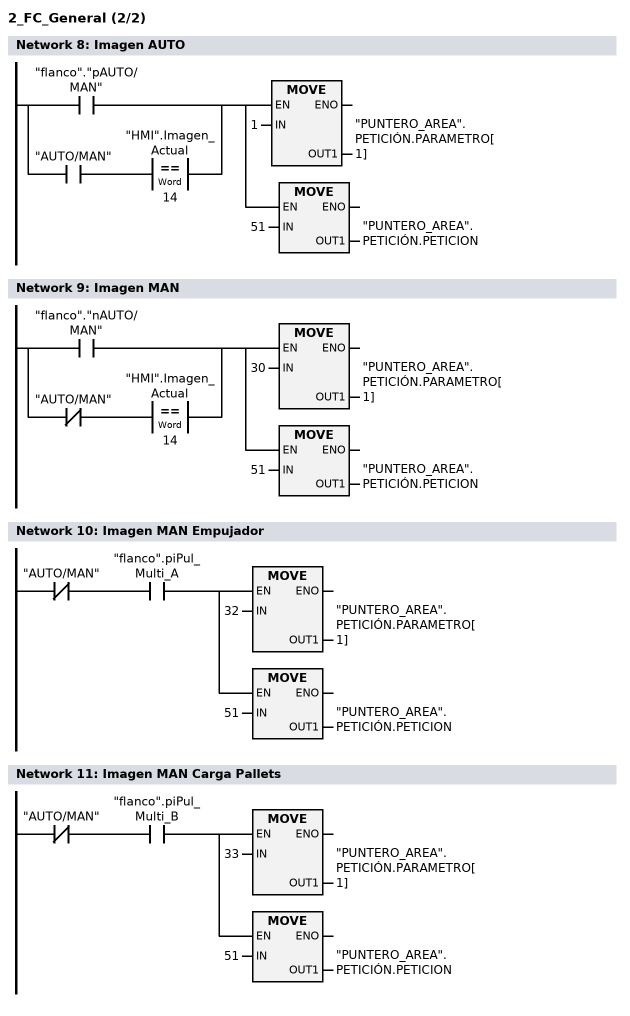
   RUNG wire#powerrail
      Contact( "flanco"."pAUTO/MAN" )
      wire#w1
      { S7_GenerateENO := "TRUE" } Move(in := 1, out1 => "PUNTERO_AREA".PETICIÓN.PARAMETRO[1])
   END_RUNG
   RUNG wire#powerrail
      Contact( "AUTO/MAN" )
      { S7_Templates := "SrcType := Word" } EQ_Contact(in1 := "HMI".Imagen_Actual, in2 := 14)
   END_RUNG wire#w1
   RUNG wire#w1
      { S7_GenerateENO := "TRUE" } Move(in := 51, out1 => "PUNTERO_AREA".PETICIÓN.PETICION)
   END_RUNG
   // the same network as SCL:
   IF "flanco"."pAUTO/MAN" OR ("AUTO/MAN" AND ("HMI".Imagen_Actual = 14)) THEN
       "PUNTERO_AREA".PETICIÓN.PARAMETRO[1] := 1;
       "PUNTERO_AREA".PETICIÓN.PETICION := 51;
   END_IF;
END_REGION

REGION Network 9: Imagen MAN
   RUNG wire#powerrail
      Contact( "flanco"."nAUTO/MAN" )
      wire#w1
      { S7_GenerateENO := "TRUE" } Move(in := 30, out1 => "PUNTERO_AREA".PETICIÓN.PARAMETRO[1])
   END_RUNG
   RUNG wire#powerrail
      I_Contact( "AUTO/MAN" )
      { S7_Templates := "SrcType := Word" } EQ_Contact(in1 := "HMI".Imagen_Actual, in2 := 14)
   END_RUNG wire#w1
   RUNG wire#w1
      { S7_GenerateENO := "TRUE" } Move(in := 51, out1 => "PUNTERO_AREA".PETICIÓN.PETICION)
   END_RUNG
   // the same network as SCL:
   IF "flanco"."nAUTO/MAN" OR (NOT "AUTO/MAN" AND ("HMI".Imagen_Actual = 14)) THEN
       "PUNTERO_AREA".PETICIÓN.PARAMETRO[1] := 30;
       "PUNTERO_AREA".PETICIÓN.PETICION := 51;
   END_IF;
END_REGION

REGION Network 10: Imagen MAN Empujador
   RUNG wire#powerrail
      I_Contact( "AUTO/MAN" )
      Contact( "flanco".piPul_Multi_A )
      wire#w1
      { S7_GenerateENO := "TRUE" } Move(in := 32, out1 => "PUNTERO_AREA".PETICIÓN.PARAMETRO[1])
   END_RUNG
   RUNG wire#w1
      { S7_GenerateENO := "TRUE" } Move(in := 51, out1 => "PUNTERO_AREA".PETICIÓN.PETICION)
   END_RUNG
   // the same network as SCL:
   IF NOT "AUTO/MAN" AND "flanco".piPul_Multi_A THEN
       "PUNTERO_AREA".PETICIÓN.PARAMETRO[1] := 32;
       "PUNTERO_AREA".PETICIÓN.PETICION := 51;
   END_IF;
END_REGION

REGION Network 11: Imagen MAN Carga Pallets
   RUNG wire#powerrail
      I_Contact( "AUTO/MAN" )
      Contact( "flanco".piPul_Multi_B )
      wire#w1
      { S7_GenerateENO := "TRUE" } Move(in := 33, out1 => "PUNTERO_AREA".PETICIÓN.PARAMETRO[1])
   END_RUNG
   RUNG wire#w1
      { S7_GenerateENO := "TRUE" } Move(in := 51, out1 => "PUNTERO_AREA".PETICIÓN.PETICION)
   END_RUNG
   // the same network as SCL:
   IF NOT "AUTO/MAN" AND "flanco".piPul_Multi_B THEN
       "PUNTERO_AREA".PETICIÓN.PARAMETRO[1] := 33;
       "PUNTERO_AREA".PETICIÓN.PETICION := 51;
   END_IF;
END_REGION
END_FUNCTION

FUNCTION "1_FC_Inv_Entradas" : Void   // FC9, LAD
{ S7_Optimized_Access := 'FALSE' }
VERSION : 0.1
BEGIN

REGION Network 1: "iiPul_DeshCargPall"
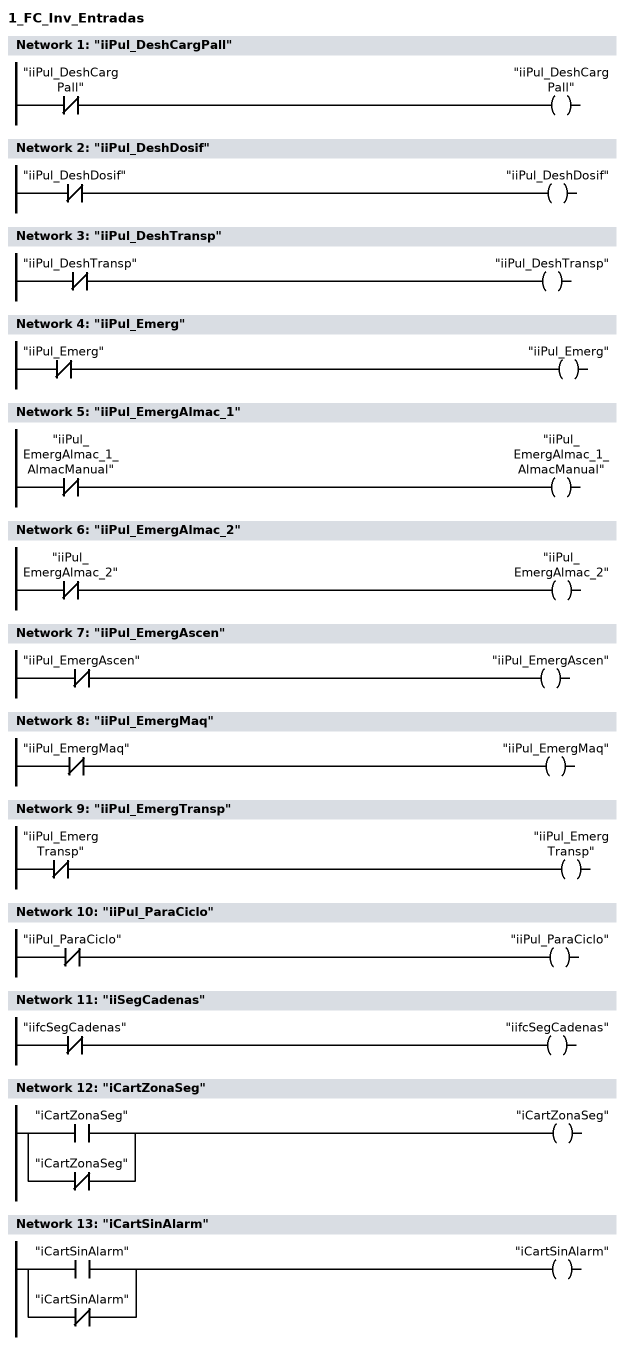
   RUNG wire#powerrail
      I_Contact( "iiPul_DeshCargPall" )
      Coil( "iiPul_DeshCargPall" )
   END_RUNG
   // the same network as SCL:
   "iiPul_DeshCargPall" := NOT "iiPul_DeshCargPall";
END_REGION

REGION Network 2: "iiPul_DeshDosif"
   RUNG wire#powerrail
      I_Contact( "iiPul_DeshDosif" )
      Coil( "iiPul_DeshDosif" )
   END_RUNG
   // the same network as SCL:
   "iiPul_DeshDosif" := NOT "iiPul_DeshDosif";
END_REGION

REGION Network 3: "iiPul_DeshTransp"
   RUNG wire#powerrail
      I_Contact( "iiPul_DeshTransp" )
      Coil( "iiPul_DeshTransp" )
   END_RUNG
   // the same network as SCL:
   "iiPul_DeshTransp" := NOT "iiPul_DeshTransp";
END_REGION

REGION Network 4: "iiPul_Emerg"
   RUNG wire#powerrail
      I_Contact( "iiPul_Emerg" )
      Coil( "iiPul_Emerg" )
   END_RUNG
   // the same network as SCL:
   "iiPul_Emerg" := NOT "iiPul_Emerg";
END_REGION

REGION Network 5: "iiPul_EmergAlmac_1"
   RUNG wire#powerrail
      I_Contact( "iiPul_EmergAlmac_1_AlmacManual" )
      Coil( "iiPul_EmergAlmac_1_AlmacManual" )
   END_RUNG
   // the same network as SCL:
   "iiPul_EmergAlmac_1_AlmacManual" := NOT "iiPul_EmergAlmac_1_AlmacManual";
END_REGION

REGION Network 6: "iiPul_EmergAlmac_2"
   RUNG wire#powerrail
      I_Contact( "iiPul_EmergAlmac_2" )
      Coil( "iiPul_EmergAlmac_2" )
   END_RUNG
   // the same network as SCL:
   "iiPul_EmergAlmac_2" := NOT "iiPul_EmergAlmac_2";
END_REGION

REGION Network 7: "iiPul_EmergAscen"
   RUNG wire#powerrail
      I_Contact( "iiPul_EmergAscen" )
      Coil( "iiPul_EmergAscen" )
   END_RUNG
   // the same network as SCL:
   "iiPul_EmergAscen" := NOT "iiPul_EmergAscen";
END_REGION

REGION Network 8: "iiPul_EmergMaq"
   RUNG wire#powerrail
      I_Contact( "iiPul_EmergMaq" )
      Coil( "iiPul_EmergMaq" )
   END_RUNG
   // the same network as SCL:
   "iiPul_EmergMaq" := NOT "iiPul_EmergMaq";
END_REGION

REGION Network 9: "iiPul_EmergTransp"
   RUNG wire#powerrail
      I_Contact( "iiPul_EmergTransp" )
      Coil( "iiPul_EmergTransp" )
   END_RUNG
   // the same network as SCL:
   "iiPul_EmergTransp" := NOT "iiPul_EmergTransp";
END_REGION

REGION Network 10: "iiPul_ParaCiclo"
   RUNG wire#powerrail
      I_Contact( "iiPul_ParaCiclo" )
      Coil( "iiPul_ParaCiclo" )
   END_RUNG
   // the same network as SCL:
   "iiPul_ParaCiclo" := NOT "iiPul_ParaCiclo";
END_REGION

REGION Network 11: "iiSegCadenas"
   RUNG wire#powerrail
      I_Contact( "iifcSegCadenas" )
      Coil( "iifcSegCadenas" )
   END_RUNG
   // the same network as SCL:
   "iifcSegCadenas" := NOT "iifcSegCadenas";
END_REGION

REGION Network 12: "iCartZonaSeg"
   RUNG wire#powerrail
      Contact( "iCartZonaSeg" )
      wire#w1
      Coil( "iCartZonaSeg" )
   END_RUNG
   RUNG wire#powerrail
      I_Contact( "iCartZonaSeg" )
   END_RUNG wire#w1
   // the same network as SCL:
   "iCartZonaSeg" := "iCartZonaSeg" OR NOT "iCartZonaSeg";
END_REGION

REGION Network 13: "iCartSinAlarm"
   RUNG wire#powerrail
      Contact( "iCartSinAlarm" )
      wire#w1
      Coil( "iCartSinAlarm" )
   END_RUNG
   RUNG wire#powerrail
      I_Contact( "iCartSinAlarm" )
   END_RUNG wire#w1
   // the same network as SCL:
   "iCartSinAlarm" := "iCartSinAlarm" OR NOT "iCartSinAlarm";
END_REGION
END_FUNCTION

FUNCTION "9_FC_Salidas" : Void   // FC10, LAD
{ S7_Optimized_Access := 'FALSE' }
VERSION : 0.1
BEGIN

REGION Network 1: "oLuz_CicloHab"
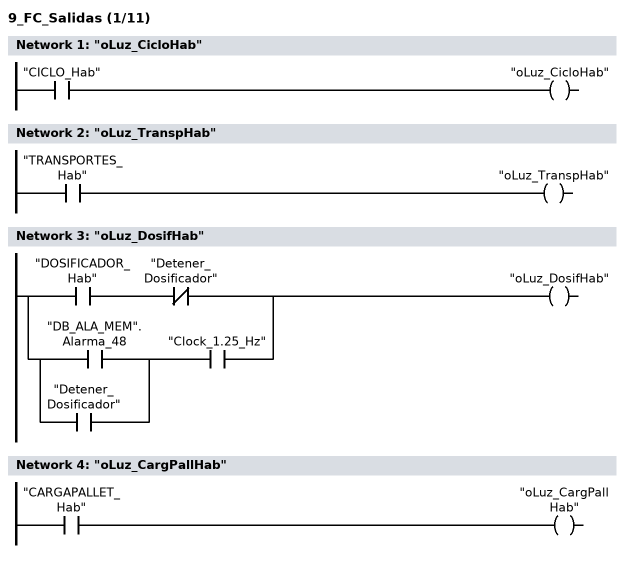
   RUNG wire#powerrail
      Contact( "CICLO_Hab" )
      Coil( "oLuz_CicloHab" )
   END_RUNG
   // the same network as SCL:
   "oLuz_CicloHab" := "CICLO_Hab";
END_REGION

REGION Network 2: "oLuz_TranspHab"
   RUNG wire#powerrail
      Contact( "TRANSPORTES_Hab" )
      Coil( "oLuz_TranspHab" )
   END_RUNG
   // the same network as SCL:
   "oLuz_TranspHab" := "TRANSPORTES_Hab";
END_REGION

REGION Network 3: "oLuz_DosifHab"
   RUNG wire#powerrail
      Contact( "DOSIFICADOR_Hab" )
      I_Contact( "Detener_Dosificador" )
      wire#w1
      Coil( "oLuz_DosifHab" )
   END_RUNG
   RUNG wire#powerrail
      Contact( "DB_ALA_MEM".Alarma_48 )
      wire#w2
      Contact( "Clock_1.25_Hz" )
   END_RUNG wire#w1
   RUNG wire#powerrail
      Contact( "Detener_Dosificador" )
   END_RUNG wire#w2
   // the same network as SCL:
   "oLuz_DosifHab" := ("DOSIFICADOR_Hab" AND NOT "Detener_Dosificador") OR (("DB_ALA_MEM".Alarma_48 OR "Detener_Dosificador") AND "Clock_1.25_Hz");
END_REGION

REGION Network 4: "oLuz_CargPallHab"
   RUNG wire#powerrail
      Contact( "CARGAPALLET_Hab" )
      Coil( "oLuz_CargPallHab" )
   END_RUNG
   // the same network as SCL:
   "oLuz_CargPallHab" := "CARGAPALLET_Hab";
END_REGION

REGION Network 5: "oLuz_Segur"
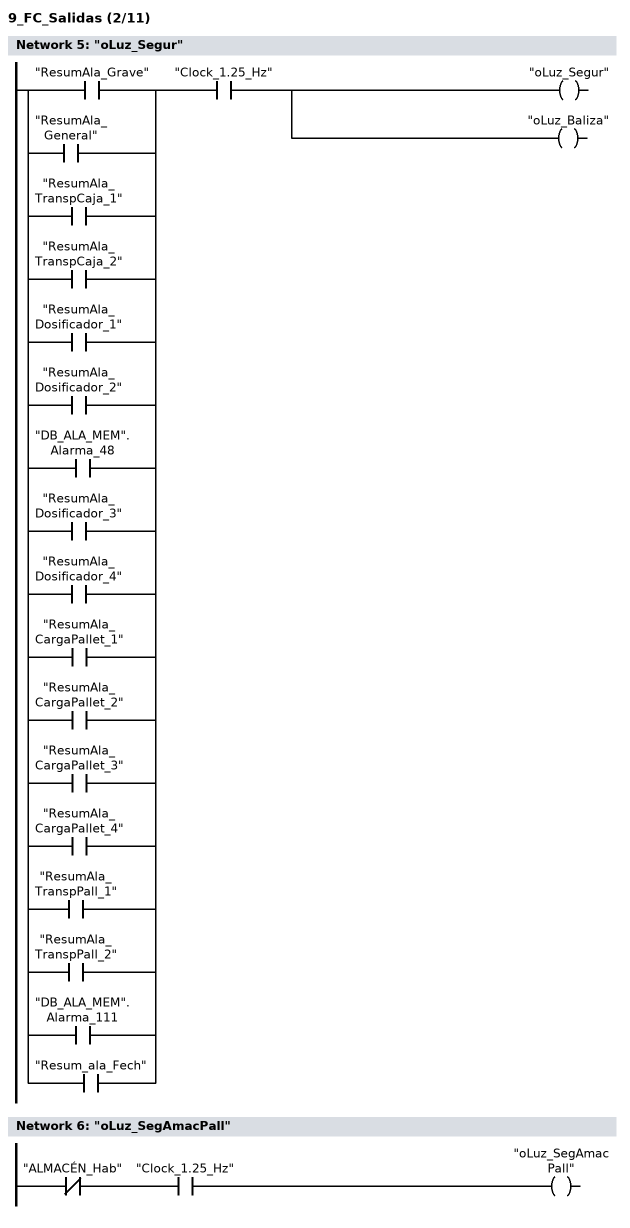
   RUNG wire#powerrail
      Contact( "ResumAla_Grave" )
      wire#w1
      Contact( "Clock_1.25_Hz" )
      wire#w2
      Coil( "oLuz_Segur" )
   END_RUNG
   RUNG wire#powerrail
      Contact( "ResumAla_General" )
   END_RUNG wire#w1
   RUNG wire#powerrail
      Contact( "ResumAla_TranspCaja_1" )
   END_RUNG wire#w1
   RUNG wire#powerrail
      Contact( "ResumAla_TranspCaja_2" )
   END_RUNG wire#w1
   RUNG wire#powerrail
      Contact( "ResumAla_Dosificador_1" )
   END_RUNG wire#w1
   RUNG wire#powerrail
      Contact( "ResumAla_Dosificador_2" )
   END_RUNG wire#w1
   RUNG wire#powerrail
      Contact( "DB_ALA_MEM".Alarma_48 )
   END_RUNG wire#w1
   RUNG wire#powerrail
      Contact( "ResumAla_Dosificador_3" )
   END_RUNG wire#w1
   RUNG wire#powerrail
      Contact( "ResumAla_Dosificador_4" )
   END_RUNG wire#w1
   RUNG wire#powerrail
      Contact( "ResumAla_CargaPallet_1" )
   END_RUNG wire#w1
   RUNG wire#powerrail
      Contact( "ResumAla_CargaPallet_2" )
   END_RUNG wire#w1
   RUNG wire#powerrail
      Contact( "ResumAla_CargaPallet_3" )
   END_RUNG wire#w1
   RUNG wire#powerrail
      Contact( "ResumAla_CargaPallet_4" )
   END_RUNG wire#w1
   RUNG wire#powerrail
      Contact( "ResumAla_TranspPall_1" )
   END_RUNG wire#w1
   RUNG wire#powerrail
      Contact( "ResumAla_TranspPall_2" )
   END_RUNG wire#w1
   RUNG wire#powerrail
      Contact( "DB_ALA_MEM".Alarma_111 )
   END_RUNG wire#w1
   RUNG wire#powerrail
      Contact( "Resum_ala_Fech" )
   END_RUNG wire#w1
   RUNG wire#w2
      Coil( "oLuz_Baliza" )
   END_RUNG
   // the same network as SCL:
   "oLuz_Segur" := ("ResumAla_Grave" OR "ResumAla_General" OR "ResumAla_TranspCaja_1" OR "ResumAla_TranspCaja_2" OR "ResumAla_Dosificador_1" OR "ResumAla_Dosificador_2" OR "DB_ALA_MEM".Alarma_48 OR "ResumAla_Dosificador_3" OR "ResumAla_Dosificador_4" OR "ResumAla_CargaPallet_1" OR "ResumAla_CargaPallet_2" OR "ResumAla_CargaPallet_3" OR "ResumAla_CargaPallet_4" OR "ResumAla_TranspPall_1" OR "ResumAla_TranspPall_2" OR "DB_ALA_MEM".Alarma_111 OR "Resum_ala_Fech") AND "Clock_1.25_Hz";
   "oLuz_Baliza" := "oLuz_Segur";
END_REGION

REGION Network 6: "oLuz_SegAmacPall"
   RUNG wire#powerrail
      I_Contact( "ALMACÉN_Hab" )
      Contact( "Clock_1.25_Hz" )
      Coil( "oLuz_SegAmacPall" )
   END_RUNG
   // the same network as SCL:
   "oLuz_SegAmacPall" := NOT "ALMACÉN_Hab" AND "Clock_1.25_Hz";
END_REGION

REGION Network 7: "oLuz_SegAscensor"
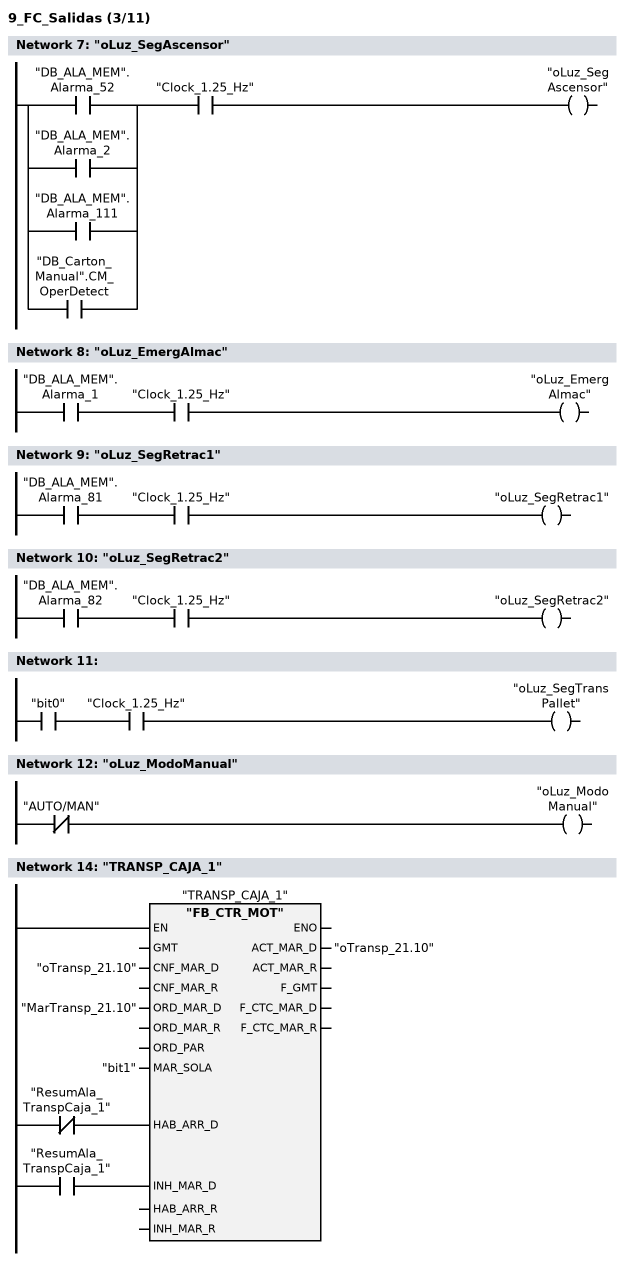
   RUNG wire#powerrail
      Contact( "DB_ALA_MEM".Alarma_52 )
      wire#w1
      Contact( "Clock_1.25_Hz" )
      Coil( "oLuz_SegAscensor" )
   END_RUNG
   RUNG wire#powerrail
      Contact( "DB_ALA_MEM".Alarma_2 )
   END_RUNG wire#w1
   RUNG wire#powerrail
      Contact( "DB_ALA_MEM".Alarma_111 )
   END_RUNG wire#w1
   RUNG wire#powerrail
      Contact( "DB_Carton_Manual".CM_OperDetect )
   END_RUNG wire#w1
   // the same network as SCL:
   "oLuz_SegAscensor" := ("DB_ALA_MEM".Alarma_52 OR "DB_ALA_MEM".Alarma_2 OR "DB_ALA_MEM".Alarma_111 OR "DB_Carton_Manual".CM_OperDetect) AND "Clock_1.25_Hz";
END_REGION

REGION Network 8: "oLuz_EmergAlmac"
   RUNG wire#powerrail
      Contact( "DB_ALA_MEM".Alarma_1 )
      Contact( "Clock_1.25_Hz" )
      Coil( "oLuz_EmergAlmac" )
   END_RUNG
   // the same network as SCL:
   "oLuz_EmergAlmac" := "DB_ALA_MEM".Alarma_1 AND "Clock_1.25_Hz";
END_REGION

REGION Network 9: "oLuz_SegRetrac1"
   RUNG wire#powerrail
      Contact( "DB_ALA_MEM".Alarma_81 )
      Contact( "Clock_1.25_Hz" )
      Coil( "oLuz_SegRetrac1" )
   END_RUNG
   // the same network as SCL:
   "oLuz_SegRetrac1" := "DB_ALA_MEM".Alarma_81 AND "Clock_1.25_Hz";
END_REGION

REGION Network 10: "oLuz_SegRetrac2"
   RUNG wire#powerrail
      Contact( "DB_ALA_MEM".Alarma_82 )
      Contact( "Clock_1.25_Hz" )
      Coil( "oLuz_SegRetrac2" )
   END_RUNG
   // the same network as SCL:
   "oLuz_SegRetrac2" := "DB_ALA_MEM".Alarma_82 AND "Clock_1.25_Hz";
END_REGION

REGION Network 11
   RUNG wire#powerrail
      Contact( "bit0" )
      Contact( "Clock_1.25_Hz" )
      Coil( "oLuz_SegTransPallet" )
   END_RUNG
   // the same network as SCL:
   "oLuz_SegTransPallet" := "bit0" AND "Clock_1.25_Hz";
END_REGION

REGION Network 12: "oLuz_ModoManual"
   RUNG wire#powerrail
      I_Contact( "AUTO/MAN" )
      Coil( "oLuz_ModoManual" )
   END_RUNG
   // the same network as SCL:
   "oLuz_ModoManual" := NOT "AUTO/MAN";
END_REGION

REGION Network 13: -------------------------------------------------- TRANSPORTES DE ENTRADA --------------------------------------------------¬
END_REGION

REGION Network 14: "TRANSP_CAJA_1"
   RUNG wire#powerrail
      "TRANSP_CAJA_1"(HAB_ARR_D := wire#w1, INH_MAR_D := wire#w2, GMT :=, CNF_MAR_D := "oTransp_21.10", CNF_MAR_R :=, ORD_MAR_D := "MarTransp_21.10", ORD_MAR_R :=, ORD_PAR :=, MAR_SOLA := "bit1", HAB_ARR_R :=, INH_MAR_R :=, ACT_MAR_D => "oTransp_21.10", ACT_MAR_R =>, F_GMT =>, F_CTC_MAR_D =>, F_CTC_MAR_R =>)
   END_RUNG
   RUNG wire#powerrail
      I_Contact( "ResumAla_TranspCaja_1" )
   END_RUNG wire#w1
   RUNG wire#powerrail
      Contact( "ResumAla_TranspCaja_1" )
   END_RUNG wire#w2
   // the same network as SCL:
   "TRANSP_CAJA_1"(CNF_MAR_D := "oTransp_21.10",   // "FB_CTR_MOT"
                   ORD_MAR_D := "MarTransp_21.10",
                   MAR_SOLA := "bit1",
                   HAB_ARR_D := NOT "ResumAla_TranspCaja_1",
                   INH_MAR_D := "ResumAla_TranspCaja_1",
                   ACT_MAR_D => "oTransp_21.10");
END_REGION

REGION Network 15: "TRANSP_CAJA_2"
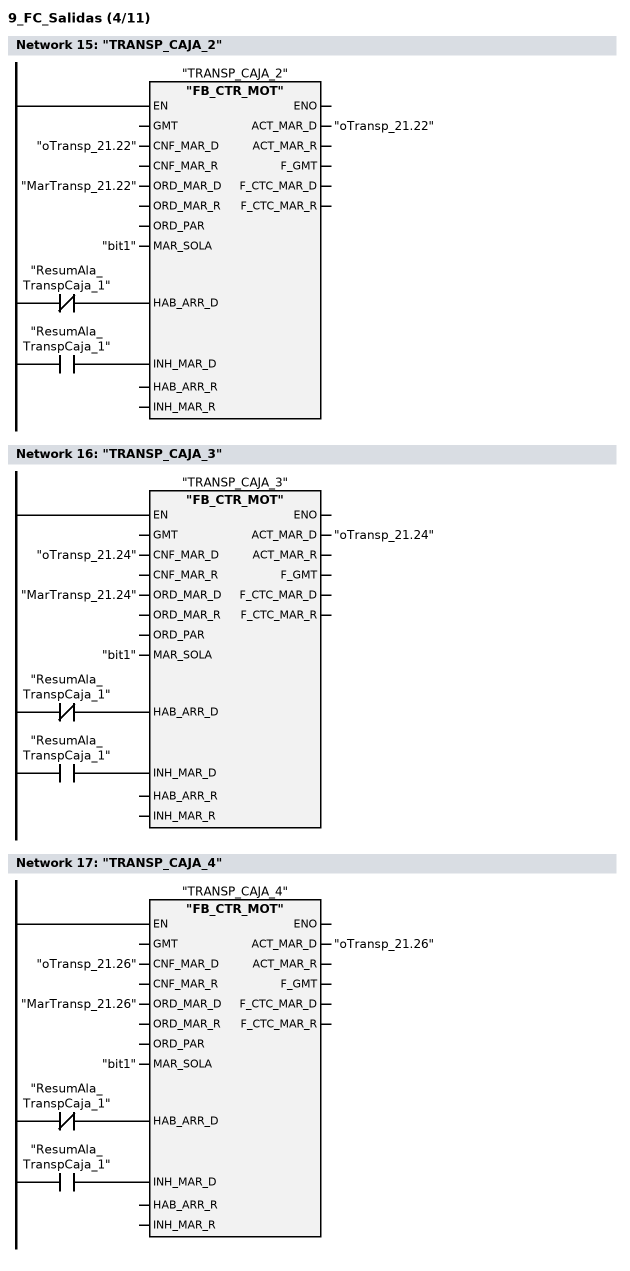
   RUNG wire#powerrail
      "TRANSP_CAJA_2"(HAB_ARR_D := wire#w1, INH_MAR_D := wire#w2, GMT :=, CNF_MAR_D := "oTransp_21.22", CNF_MAR_R :=, ORD_MAR_D := "MarTransp_21.22", ORD_MAR_R :=, ORD_PAR :=, MAR_SOLA := "bit1", HAB_ARR_R :=, INH_MAR_R :=, ACT_MAR_D => "oTransp_21.22", ACT_MAR_R =>, F_GMT =>, F_CTC_MAR_D =>, F_CTC_MAR_R =>)
   END_RUNG
   RUNG wire#powerrail
      I_Contact( "ResumAla_TranspCaja_1" )
   END_RUNG wire#w1
   RUNG wire#powerrail
      Contact( "ResumAla_TranspCaja_1" )
   END_RUNG wire#w2
   // the same network as SCL:
   "TRANSP_CAJA_2"(CNF_MAR_D := "oTransp_21.22",   // "FB_CTR_MOT"
                   ORD_MAR_D := "MarTransp_21.22",
                   MAR_SOLA := "bit1",
                   HAB_ARR_D := NOT "ResumAla_TranspCaja_1",
                   INH_MAR_D := "ResumAla_TranspCaja_1",
                   ACT_MAR_D => "oTransp_21.22");
END_REGION

REGION Network 16: "TRANSP_CAJA_3"
   RUNG wire#powerrail
      "TRANSP_CAJA_3"(HAB_ARR_D := wire#w1, INH_MAR_D := wire#w2, GMT :=, CNF_MAR_D := "oTransp_21.24", CNF_MAR_R :=, ORD_MAR_D := "MarTransp_21.24", ORD_MAR_R :=, ORD_PAR :=, MAR_SOLA := "bit1", HAB_ARR_R :=, INH_MAR_R :=, ACT_MAR_D => "oTransp_21.24", ACT_MAR_R =>, F_GMT =>, F_CTC_MAR_D =>, F_CTC_MAR_R =>)
   END_RUNG
   RUNG wire#powerrail
      I_Contact( "ResumAla_TranspCaja_1" )
   END_RUNG wire#w1
   RUNG wire#powerrail
      Contact( "ResumAla_TranspCaja_1" )
   END_RUNG wire#w2
   // the same network as SCL:
   "TRANSP_CAJA_3"(CNF_MAR_D := "oTransp_21.24",   // "FB_CTR_MOT"
                   ORD_MAR_D := "MarTransp_21.24",
                   MAR_SOLA := "bit1",
                   HAB_ARR_D := NOT "ResumAla_TranspCaja_1",
                   INH_MAR_D := "ResumAla_TranspCaja_1",
                   ACT_MAR_D => "oTransp_21.24");
END_REGION

REGION Network 17: "TRANSP_CAJA_4"
   RUNG wire#powerrail
      "TRANSP_CAJA_4"(HAB_ARR_D := wire#w1, INH_MAR_D := wire#w2, GMT :=, CNF_MAR_D := "oTransp_21.26", CNF_MAR_R :=, ORD_MAR_D := "MarTransp_21.26", ORD_MAR_R :=, ORD_PAR :=, MAR_SOLA := "bit1", HAB_ARR_R :=, INH_MAR_R :=, ACT_MAR_D => "oTransp_21.26", ACT_MAR_R =>, F_GMT =>, F_CTC_MAR_D =>, F_CTC_MAR_R =>)
   END_RUNG
   RUNG wire#powerrail
      I_Contact( "ResumAla_TranspCaja_1" )
   END_RUNG wire#w1
   RUNG wire#powerrail
      Contact( "ResumAla_TranspCaja_1" )
   END_RUNG wire#w2
   // the same network as SCL:
   "TRANSP_CAJA_4"(CNF_MAR_D := "oTransp_21.26",   // "FB_CTR_MOT"
                   ORD_MAR_D := "MarTransp_21.26",
                   MAR_SOLA := "bit1",
                   HAB_ARR_D := NOT "ResumAla_TranspCaja_1",
                   INH_MAR_D := "ResumAla_TranspCaja_1",
                   ACT_MAR_D => "oTransp_21.26");
END_REGION

REGION Network 18: -------------------------------------------------------------- DOSIFICADOR --------------------------------------------------------------¬
END_REGION

REGION Network 19: "VARIADOR_DOSIFICADOR"
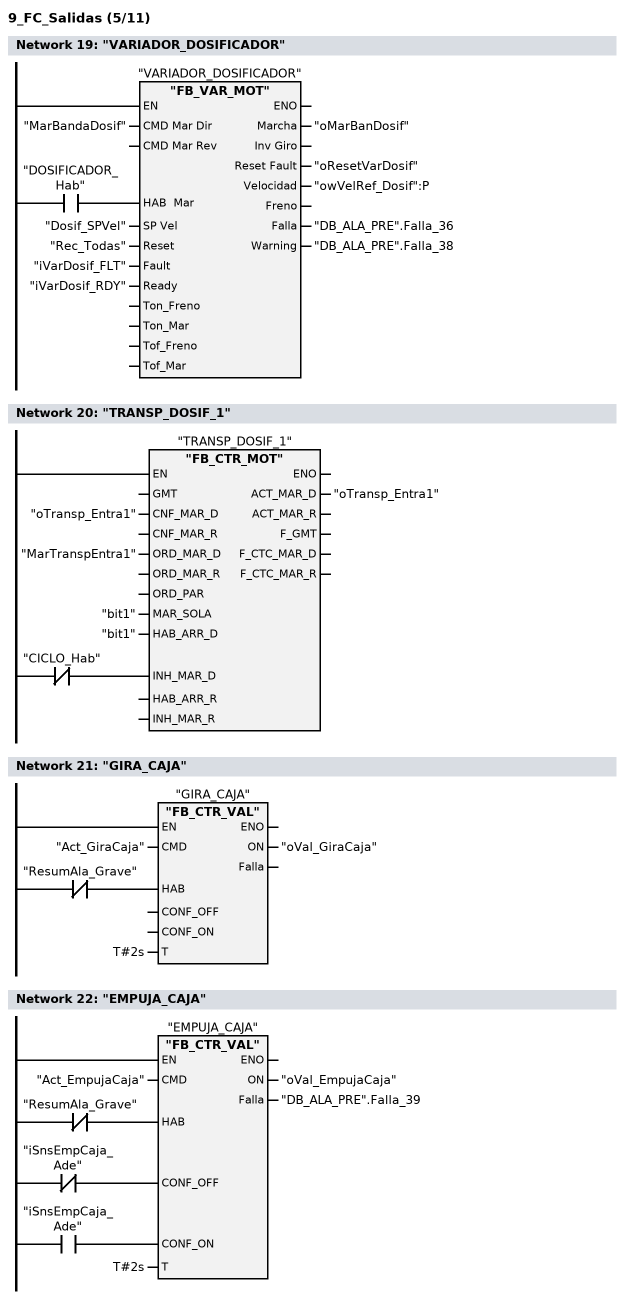
   RUNG wire#powerrail
      "VARIADOR_DOSIFICADOR"("HAB  Mar" := wire#w1, "CMD Mar Dir" := "MarBandaDosif", "CMD Mar Rev" :=, "SP Vel" := "Dosif_SPVel", Reset := "Rec_Todas", Fault := "iVarDosif_FLT", Ready := "iVarDosif_RDY", Ton_Freno :=, Ton_Mar :=, Tof_Freno :=, Tof_Mar :=, Marcha => "oMarBanDosif", "Inv Giro" =>, "Reset Fault" => "oResetVarDosif", Velocidad => "owVelRef_Dosif":P, Freno =>, Falla => "DB_ALA_PRE".Falla_36, Warning => "DB_ALA_PRE".Falla_38)
   END_RUNG
   RUNG wire#powerrail
      Contact( "DOSIFICADOR_Hab" )
   END_RUNG wire#w1
   // the same network as SCL:
   "VARIADOR_DOSIFICADOR"("CMD Mar Dir" := "MarBandaDosif",   // "FB_VAR_MOT"
                          "HAB  Mar" := "DOSIFICADOR_Hab",
                          "SP Vel" := "Dosif_SPVel",
                          Reset := "Rec_Todas",
                          Fault := "iVarDosif_FLT",
                          Ready := "iVarDosif_RDY",
                          Marcha => "oMarBanDosif",
                          "Reset Fault" => "oResetVarDosif",
                          Velocidad => "owVelRef_Dosif":P,
                          Falla => "DB_ALA_PRE".Falla_36,
                          Warning => "DB_ALA_PRE".Falla_38);
END_REGION

REGION Network 20: "TRANSP_DOSIF_1"
   RUNG wire#powerrail
      "TRANSP_DOSIF_1"(INH_MAR_D := wire#w1, GMT :=, CNF_MAR_D := "oTransp_Entra1", CNF_MAR_R :=, ORD_MAR_D := "MarTranspEntra1", ORD_MAR_R :=, ORD_PAR :=, MAR_SOLA := "bit1", HAB_ARR_D := "bit1", HAB_ARR_R :=, INH_MAR_R :=, ACT_MAR_D => "oTransp_Entra1", ACT_MAR_R =>, F_GMT =>, F_CTC_MAR_D =>, F_CTC_MAR_R =>)
   END_RUNG
   RUNG wire#powerrail
      I_Contact( "CICLO_Hab" )
   END_RUNG wire#w1
   // the same network as SCL:
   "TRANSP_DOSIF_1"(CNF_MAR_D := "oTransp_Entra1",   // "FB_CTR_MOT"
                    ORD_MAR_D := "MarTranspEntra1",
                    MAR_SOLA := "bit1",
                    HAB_ARR_D := "bit1",
                    INH_MAR_D := NOT "CICLO_Hab",
                    ACT_MAR_D => "oTransp_Entra1");
END_REGION

REGION Network 21: "GIRA_CAJA"
   RUNG wire#powerrail
      "GIRA_CAJA"(HAB := wire#w1, CMD := "Act_GiraCaja", CONF_OFF :=, CONF_ON :=, T := T#2s, ON => "oVal_GiraCaja", Falla =>)
   END_RUNG
   RUNG wire#powerrail
      I_Contact( "ResumAla_Grave" )
   END_RUNG wire#w1
   // the same network as SCL:
   "GIRA_CAJA"(CMD := "Act_GiraCaja", HAB := NOT "ResumAla_Grave", T := T#2s, ON => "oVal_GiraCaja");   // "FB_CTR_VAL"
END_REGION

REGION Network 22: "EMPUJA_CAJA"
   RUNG wire#powerrail
      "EMPUJA_CAJA"(HAB := wire#w1, CONF_OFF := wire#w2, CONF_ON := wire#w3, CMD := "Act_EmpujaCaja", T := T#2s, ON => "oVal_EmpujaCaja", Falla => "DB_ALA_PRE".Falla_39)
   END_RUNG
   RUNG wire#powerrail
      I_Contact( "ResumAla_Grave" )
   END_RUNG wire#w1
   RUNG wire#powerrail
      I_Contact( "iSnsEmpCaja_Ade" )
   END_RUNG wire#w2
   RUNG wire#powerrail
      Contact( "iSnsEmpCaja_Ade" )
   END_RUNG wire#w3
   // the same network as SCL:
   "EMPUJA_CAJA"(CMD := "Act_EmpujaCaja",   // "FB_CTR_VAL"
                 HAB := NOT "ResumAla_Grave",
                 CONF_OFF := NOT "iSnsEmpCaja_Ade",
                 CONF_ON := "iSnsEmpCaja_Ade",
                 T := T#2s,
                 ON => "oVal_EmpujaCaja",
                 Falla => "DB_ALA_PRE".Falla_39);
END_REGION

REGION Network 23: "STOP_CAJA"
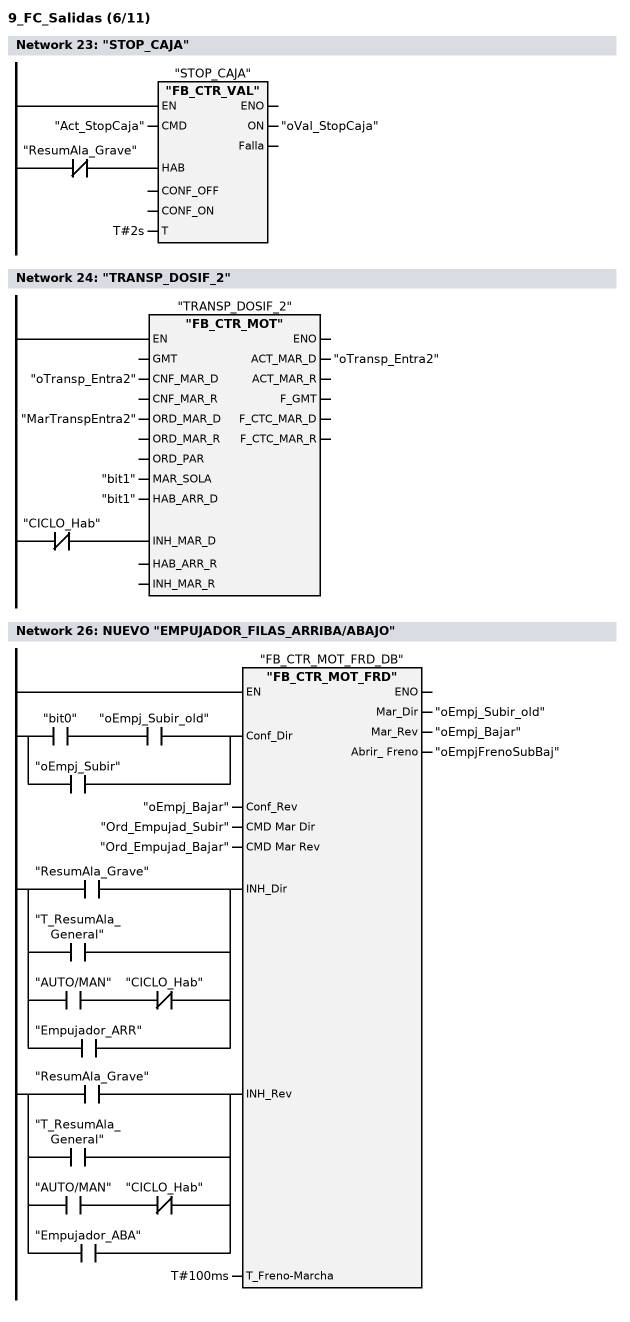
   RUNG wire#powerrail
      "STOP_CAJA"(HAB := wire#w1, CMD := "Act_StopCaja", CONF_OFF :=, CONF_ON :=, T := T#2s, ON => "oVal_StopCaja", Falla =>)
   END_RUNG
   RUNG wire#powerrail
      I_Contact( "ResumAla_Grave" )
   END_RUNG wire#w1
   // the same network as SCL:
   "STOP_CAJA"(CMD := "Act_StopCaja", HAB := NOT "ResumAla_Grave", T := T#2s, ON => "oVal_StopCaja");   // "FB_CTR_VAL"
END_REGION

REGION Network 24: "TRANSP_DOSIF_2"
   RUNG wire#powerrail
      "TRANSP_DOSIF_2"(INH_MAR_D := wire#w1, GMT :=, CNF_MAR_D := "oTransp_Entra2", CNF_MAR_R :=, ORD_MAR_D := "MarTranspEntra2", ORD_MAR_R :=, ORD_PAR :=, MAR_SOLA := "bit1", HAB_ARR_D := "bit1", HAB_ARR_R :=, INH_MAR_R :=, ACT_MAR_D => "oTransp_Entra2", ACT_MAR_R =>, F_GMT =>, F_CTC_MAR_D =>, F_CTC_MAR_R =>)
   END_RUNG
   RUNG wire#powerrail
      I_Contact( "CICLO_Hab" )
   END_RUNG wire#w1
   // the same network as SCL:
   "TRANSP_DOSIF_2"(CNF_MAR_D := "oTransp_Entra2",   // "FB_CTR_MOT"
                    ORD_MAR_D := "MarTranspEntra2",
                    MAR_SOLA := "bit1",
                    HAB_ARR_D := "bit1",
                    INH_MAR_D := NOT "CICLO_Hab",
                    ACT_MAR_D => "oTransp_Entra2");
END_REGION

REGION Network 25: ------------------------------------------------------------------ EMPUJADOR ------------------------------------------------------------------¬
END_REGION

REGION Network 26: NUEVO "EMPUJADOR_FILAS_ARRIBA/ABAJO"
   RUNG wire#powerrail
      "FB_CTR_MOT_FRD_DB"(Conf_Dir := wire#w1, INH_Dir := wire#w2, INH_Rev := wire#w3, Conf_Rev := "oEmpj_Bajar", "CMD Mar Dir" := "Ord_Empujad_Subir", "CMD Mar Rev" := "Ord_Empujad_Bajar", "T_Freno-Marcha" := T#100ms, Mar_Dir => "oEmpj_Subir_old", Mar_Rev => "oEmpj_Bajar", "Abrir_ Freno" => "oEmpjFrenoSubBaj")
   END_RUNG
   RUNG wire#powerrail
      Contact( "bit0" )
      Contact( "oEmpj_Subir_old" )
   END_RUNG wire#w1
   RUNG wire#powerrail
      Contact( "oEmpj_Subir" )
   END_RUNG wire#w1
   RUNG wire#powerrail
      Contact( "ResumAla_Grave" )
   END_RUNG wire#w2
   RUNG wire#powerrail
      Contact( "T_ResumAla_General" )
   END_RUNG wire#w2
   RUNG wire#powerrail
      Contact( "AUTO/MAN" )
      I_Contact( "CICLO_Hab" )
   END_RUNG wire#w2
   RUNG wire#powerrail
      Contact( "Empujador_ARR" )
   END_RUNG wire#w2
   RUNG wire#powerrail
      Contact( "ResumAla_Grave" )
   END_RUNG wire#w3
   RUNG wire#powerrail
      Contact( "T_ResumAla_General" )
   END_RUNG wire#w3
   RUNG wire#powerrail
      Contact( "AUTO/MAN" )
      I_Contact( "CICLO_Hab" )
   END_RUNG wire#w3
   RUNG wire#powerrail
      Contact( "Empujador_ABA" )
   END_RUNG wire#w3
   // the same network as SCL:
   "FB_CTR_MOT_FRD_DB"(Conf_Dir := ("bit0" AND "oEmpj_Subir_old") OR "oEmpj_Subir",   // "FB_CTR_MOT_FRD"
                       Conf_Rev := "oEmpj_Bajar",
                       "CMD Mar Dir" := "Ord_Empujad_Subir",
                       "CMD Mar Rev" := "Ord_Empujad_Bajar",
                       INH_Dir := "ResumAla_Grave" OR "T_ResumAla_General" OR ("AUTO/MAN" AND NOT "CICLO_Hab") OR "Empujador_ARR",
                       INH_Rev := "ResumAla_Grave" OR "T_ResumAla_General" OR ("AUTO/MAN" AND NOT "CICLO_Hab") OR "Empujador_ABA",
                       "T_Freno-Marcha" := T#100ms,
                       Mar_Dir => "oEmpj_Subir_old",
                       Mar_Rev => "oEmpj_Bajar",
                       "Abrir_ Freno" => "oEmpjFrenoSubBaj");
END_REGION

REGION Network 27: "EMPUJADOR_FILAS_ADELANTE/ATRÁS"
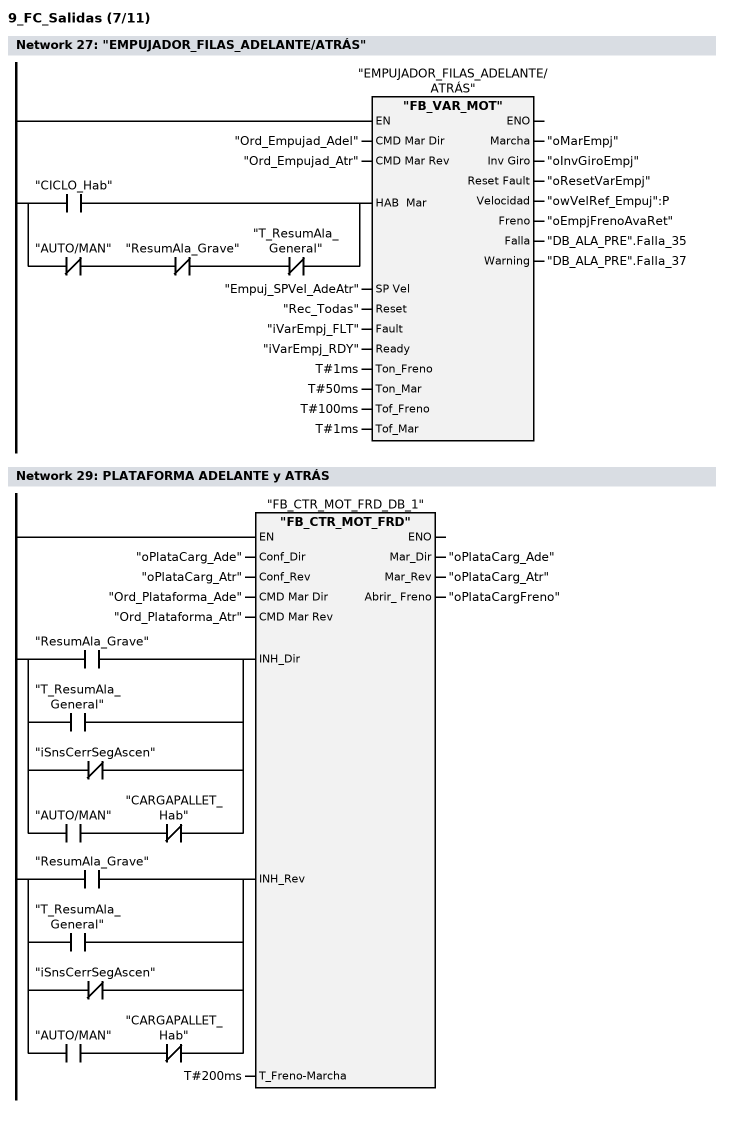
   RUNG wire#powerrail
      "EMPUJADOR_FILAS_ADELANTE/ATRÁS"("HAB  Mar" := wire#w1, "CMD Mar Dir" := "Ord_Empujad_Adel", "CMD Mar Rev" := "Ord_Empujad_Atr", "SP Vel" := "Empuj_SPVel_AdeAtr", Reset := "Rec_Todas", Fault := "iVarEmpj_FLT", Ready := "iVarEmpj_RDY", Ton_Freno := T#1ms, Ton_Mar := T#50ms, Tof_Freno := T#100ms, Tof_Mar := T#1ms, Marcha => "oMarEmpj", "Inv Giro" => "oInvGiroEmpj", "Reset Fault" => "oResetVarEmpj", Velocidad => "owVelRef_Empuj":P, Freno => "oEmpjFrenoAvaRet", Falla => "DB_ALA_PRE".Falla_35, Warning => "DB_ALA_PRE".Falla_37)
   END_RUNG
   RUNG wire#powerrail
      Contact( "CICLO_Hab" )
   END_RUNG wire#w1
   RUNG wire#powerrail
      I_Contact( "AUTO/MAN" )
      I_Contact( "ResumAla_Grave" )
      I_Contact( "T_ResumAla_General" )
   END_RUNG wire#w1
   // the same network as SCL:
   "EMPUJADOR_FILAS_ADELANTE/ATRÁS"("CMD Mar Dir" := "Ord_Empujad_Adel",   // "FB_VAR_MOT"
                           "CMD Mar Rev" := "Ord_Empujad_Atr",
                           "HAB  Mar" := "CICLO_Hab" OR (NOT "AUTO/MAN" AND NOT "ResumAla_Grave" AND NOT "T_ResumAla_General"),
                           "SP Vel" := "Empuj_SPVel_AdeAtr",
                           Reset := "Rec_Todas",
                           Fault := "iVarEmpj_FLT",
                           Ready := "iVarEmpj_RDY",
                           Ton_Freno := T#1ms,
                           Ton_Mar := T#50ms,
                           Tof_Freno := T#100ms,
                           Tof_Mar := T#1ms,
                           Marcha => "oMarEmpj",
                           "Inv Giro" => "oInvGiroEmpj",
                           "Reset Fault" => "oResetVarEmpj",
                           Velocidad => "owVelRef_Empuj":P,
                           Freno => "oEmpjFrenoAvaRet",
                           Falla => "DB_ALA_PRE".Falla_35,
                           Warning => "DB_ALA_PRE".Falla_37);
END_REGION

REGION Network 28: ----------------------------------------------------------------- CARGA DE PALLETS -----------------------------------------------------------------¬
END_REGION
